
REGION Network 78: Sin requerimiento compresor 5
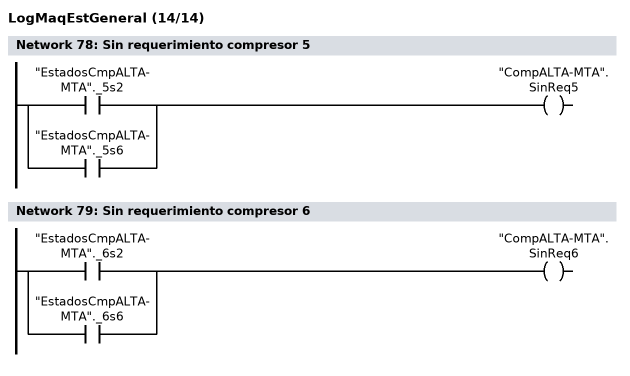
   RUNG wire#powerrail
      Contact( "EstadosCmpALTA-MTA"._5s2 )
      wire#w1
      Coil( "CompALTA-MTA".SinReq5 )
   END_RUNG
   RUNG wire#powerrail
      Contact( "EstadosCmpALTA-MTA"._5s6 )
   END_RUNG wire#w1
   // the same network as SCL:
   "CompALTA-MTA".SinReq5 := "EstadosCmpALTA-MTA"._5s2 OR "EstadosCmpALTA-MTA"._5s6;
END_REGION

REGION Network 79: Sin requerimiento compresor 6
   RUNG wire#powerrail
      Contact( "EstadosCmpALTA-MTA"._6s2 )
      wire#w1
      Coil( "CompALTA-MTA".SinReq6 )
   END_RUNG
   RUNG wire#powerrail
      Contact( "EstadosCmpALTA-MTA"._6s6 )
   END_RUNG wire#w1
   // the same network as SCL:
   "CompALTA-MTA".SinReq6 := "EstadosCmpALTA-MTA"._6s2 OR "EstadosCmpALTA-MTA"._6s6;
END_REGION
END_FUNCTION

FUNCTION "CalcEst1" : Void   // FC36, LAD
{ S7_Optimized_Access := 'FALSE' }
VERSION : 0.1
   VAR_TEMP   // added for the SCL form of the ladder/FBD networks
      _w1 : Bool;
   END_VAR
BEGIN

REGION Network 1
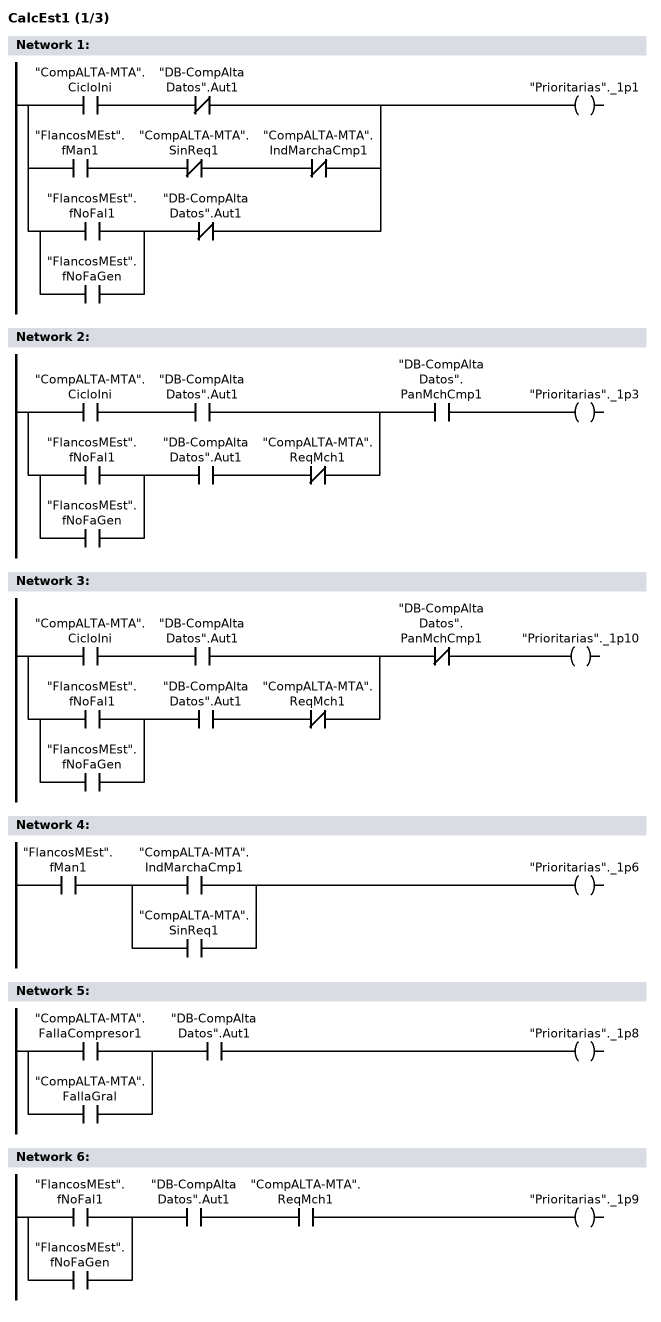
   RUNG wire#powerrail
      Contact( "CompALTA-MTA".CicloIni )
      I_Contact( "DB-CompAltaDatos".Aut1 )
      wire#w1
      Coil( "Prioritarias"._1p1 )
   END_RUNG
   RUNG wire#powerrail
      Contact( "FlancosMEst".fMan1 )
      I_Contact( "CompALTA-MTA".SinReq1 )
      I_Contact( "CompALTA-MTA".IndMarchaCmp1 )
   END_RUNG wire#w1
   RUNG wire#powerrail
      Contact( "FlancosMEst".fNoFal1 )
      wire#w2
      I_Contact( "DB-CompAltaDatos".Aut1 )
   END_RUNG wire#w1
   RUNG wire#powerrail
      Contact( "FlancosMEst".fNoFaGen )
   END_RUNG wire#w2
   // the same network as SCL:
   "Prioritarias"._1p1 := ("CompALTA-MTA".CicloIni AND NOT "DB-CompAltaDatos".Aut1) OR ("FlancosMEst".fMan1 AND NOT "CompALTA-MTA".SinReq1 AND NOT "CompALTA-MTA".IndMarchaCmp1) OR (("FlancosMEst".fNoFal1 OR "FlancosMEst".fNoFaGen) AND NOT "DB-CompAltaDatos".Aut1);
END_REGION

REGION Network 2
   RUNG wire#powerrail
      Contact( "CompALTA-MTA".CicloIni )
      Contact( "DB-CompAltaDatos".Aut1 )
      wire#w1
      Contact( "DB-CompAltaDatos".PanMchCmp1 )
      Coil( "Prioritarias"._1p3 )
   END_RUNG
   RUNG wire#powerrail
      Contact( "FlancosMEst".fNoFal1 )
      wire#w2
      Contact( "DB-CompAltaDatos".Aut1 )
      I_Contact( "CompALTA-MTA".ReqMch1 )
   END_RUNG wire#w1
   RUNG wire#powerrail
      Contact( "FlancosMEst".fNoFaGen )
   END_RUNG wire#w2
   // the same network as SCL:
   "Prioritarias"._1p3 := (("CompALTA-MTA".CicloIni AND "DB-CompAltaDatos".Aut1) OR (("FlancosMEst".fNoFal1 OR "FlancosMEst".fNoFaGen) AND "DB-CompAltaDatos".Aut1 AND NOT "CompALTA-MTA".ReqMch1)) AND "DB-CompAltaDatos".PanMchCmp1;
END_REGION

REGION Network 3
   RUNG wire#powerrail
      Contact( "CompALTA-MTA".CicloIni )
      Contact( "DB-CompAltaDatos".Aut1 )
      wire#w1
      I_Contact( "DB-CompAltaDatos".PanMchCmp1 )
      Coil( "Prioritarias"._1p10 )
   END_RUNG
   RUNG wire#powerrail
      Contact( "FlancosMEst".fNoFal1 )
      wire#w2
      Contact( "DB-CompAltaDatos".Aut1 )
      I_Contact( "CompALTA-MTA".ReqMch1 )
   END_RUNG wire#w1
   RUNG wire#powerrail
      Contact( "FlancosMEst".fNoFaGen )
   END_RUNG wire#w2
   // the same network as SCL:
   "Prioritarias"._1p10 := (("CompALTA-MTA".CicloIni AND "DB-CompAltaDatos".Aut1) OR (("FlancosMEst".fNoFal1 OR "FlancosMEst".fNoFaGen) AND "DB-CompAltaDatos".Aut1 AND NOT "CompALTA-MTA".ReqMch1)) AND NOT "DB-CompAltaDatos".PanMchCmp1;
END_REGION

REGION Network 4
   RUNG wire#powerrail
      Contact( "FlancosMEst".fMan1 )
      wire#w1
      Contact( "CompALTA-MTA".IndMarchaCmp1 )
      wire#w2
      Coil( "Prioritarias"._1p6 )
   END_RUNG
   RUNG wire#w1
      Contact( "CompALTA-MTA".SinReq1 )
   END_RUNG wire#w2
   // the same network as SCL:
   "Prioritarias"._1p6 := "FlancosMEst".fMan1 AND ("CompALTA-MTA".IndMarchaCmp1 OR "CompALTA-MTA".SinReq1);
END_REGION

REGION Network 5
   RUNG wire#powerrail
      Contact( "CompALTA-MTA".FallaCompresor1 )
      wire#w1
      Contact( "DB-CompAltaDatos".Aut1 )
      Coil( "Prioritarias"._1p8 )
   END_RUNG
   RUNG wire#powerrail
      Contact( "CompALTA-MTA".FallaGral )
   END_RUNG wire#w1
   // the same network as SCL:
   "Prioritarias"._1p8 := ("CompALTA-MTA".FallaCompresor1 OR "CompALTA-MTA".FallaGral) AND "DB-CompAltaDatos".Aut1;
END_REGION

REGION Network 6
   RUNG wire#powerrail
      Contact( "FlancosMEst".fNoFal1 )
      wire#w1
      Contact( "DB-CompAltaDatos".Aut1 )
      Contact( "CompALTA-MTA".ReqMch1 )
      Coil( "Prioritarias"._1p9 )
   END_RUNG
   RUNG wire#powerrail
      Contact( "FlancosMEst".fNoFaGen )
   END_RUNG wire#w1
   // the same network as SCL:
   "Prioritarias"._1p9 := ("FlancosMEst".fNoFal1 OR "FlancosMEst".fNoFaGen) AND "DB-CompAltaDatos".Aut1 AND "CompALTA-MTA".ReqMch1;
END_REGION

REGION Network 7
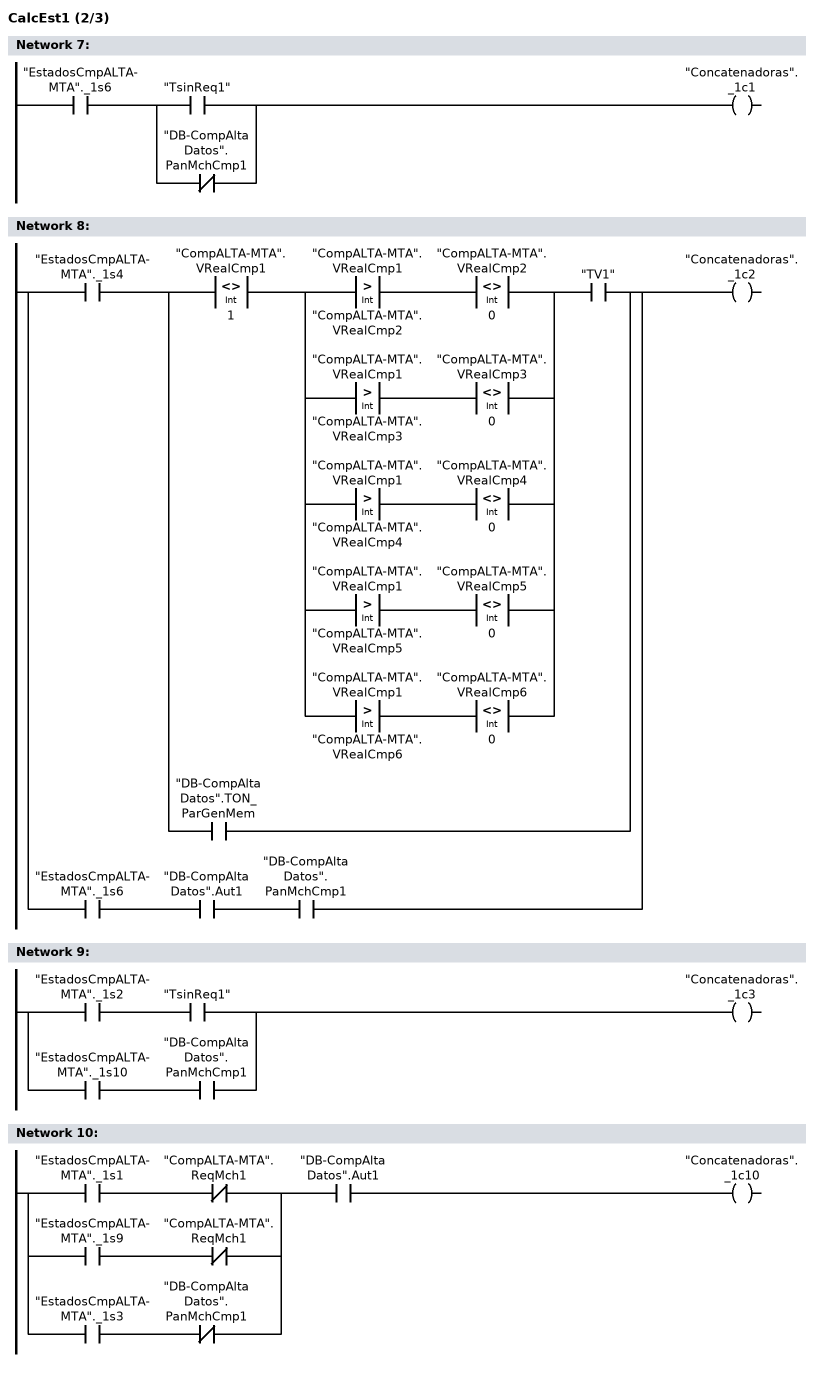
   RUNG wire#powerrail
      Contact( "EstadosCmpALTA-MTA"._1s6 )
      wire#w1
      Contact( "TsinReq1" )
      wire#w2
      Coil( "Concatenadoras"._1c1 )
   END_RUNG
   RUNG wire#w1
      I_Contact( "DB-CompAltaDatos".PanMchCmp1 )
   END_RUNG wire#w2
   // the same network as SCL:
   "Concatenadoras"._1c1 := "EstadosCmpALTA-MTA"._1s6 AND ("TsinReq1" OR NOT "DB-CompAltaDatos".PanMchCmp1);
END_REGION

REGION Network 8
   RUNG wire#powerrail
      Contact( "EstadosCmpALTA-MTA"._1s4 )
      wire#w1
      { S7_Templates := "SrcType := Int" } NE_Contact(in1 := "CompALTA-MTA".VRealCmp1, in2 := 1)
      wire#w2
      { S7_Templates := "SrcType := Int" } GT_Contact(in1 := "CompALTA-MTA".VRealCmp1, in2 := "CompALTA-MTA".VRealCmp2)
      { S7_Templates := "SrcType := Int" } NE_Contact(in1 := "CompALTA-MTA".VRealCmp2, in2 := 0)
      wire#w3
      Contact( "TV1" )
      wire#w4
      Coil( "Concatenadoras"._1c2 )
   END_RUNG
   RUNG wire#w2
      { S7_Templates := "SrcType := Int" } GT_Contact(in1 := "CompALTA-MTA".VRealCmp1, in2 := "CompALTA-MTA".VRealCmp3)
      { S7_Templates := "SrcType := Int" } NE_Contact(in1 := "CompALTA-MTA".VRealCmp3, in2 := 0)
   END_RUNG wire#w3
   RUNG wire#w2
      { S7_Templates := "SrcType := Int" } GT_Contact(in1 := "CompALTA-MTA".VRealCmp1, in2 := "CompALTA-MTA".VRealCmp4)
      { S7_Templates := "SrcType := Int" } NE_Contact(in1 := "CompALTA-MTA".VRealCmp4, in2 := 0)
   END_RUNG wire#w3
   RUNG wire#w2
      { S7_Templates := "SrcType := Int" } GT_Contact(in1 := "CompALTA-MTA".VRealCmp1, in2 := "CompALTA-MTA".VRealCmp5)
      { S7_Templates := "SrcType := Int" } NE_Contact(in1 := "CompALTA-MTA".VRealCmp5, in2 := 0)
   END_RUNG wire#w3
   RUNG wire#w2
      { S7_Templates := "SrcType := Int" } GT_Contact(in1 := "CompALTA-MTA".VRealCmp1, in2 := "CompALTA-MTA".VRealCmp6)
      { S7_Templates := "SrcType := Int" } NE_Contact(in1 := "CompALTA-MTA".VRealCmp6, in2 := 0)
   END_RUNG wire#w3
   RUNG wire#w1
      Contact( "DB-CompAltaDatos".TON_ParGenMem )
   END_RUNG wire#w4
   RUNG wire#powerrail
      Contact( "EstadosCmpALTA-MTA"._1s6 )
      Contact( "DB-CompAltaDatos".Aut1 )
      Contact( "DB-CompAltaDatos".PanMchCmp1 )
   END_RUNG wire#w4
   // the same network as SCL:
   "Concatenadoras"._1c2 := ("EstadosCmpALTA-MTA"._1s4 AND ((("CompALTA-MTA".VRealCmp1 <> 1) AND ((("CompALTA-MTA".VRealCmp1 > "CompALTA-MTA".VRealCmp2) AND ("CompALTA-MTA".VRealCmp2 <> 0)) OR (("CompALTA-MTA".VRealCmp1 > "CompALTA-MTA".VRealCmp3) AND ("CompALTA-MTA".VRealCmp3 <> 0)) OR (("CompALTA-MTA".VRealCmp1 > "CompALTA-MTA".VRealCmp4) AND ("CompALTA-MTA".VRealCmp4 <> 0)) OR (("CompALTA-MTA".VRealCmp1 > "CompALTA-MTA".VRealCmp5) AND ("CompALTA-MTA".VRealCmp5 <> 0)) OR (("CompALTA-MTA".VRealCmp1 > "CompALTA-MTA".VRealCmp6) AND ("CompALTA-MTA".VRealCmp6 <> 0))) AND "TV1") OR "DB-CompAltaDatos".TON_ParGenMem)) OR ("EstadosCmpALTA-MTA"._1s6 AND "DB-CompAltaDatos".Aut1 AND "DB-CompAltaDatos".PanMchCmp1);
END_REGION

REGION Network 9
   RUNG wire#powerrail
      Contact( "EstadosCmpALTA-MTA"._1s2 )
      Contact( "TsinReq1" )
      wire#w1
      Coil( "Concatenadoras"._1c3 )
   END_RUNG
   RUNG wire#powerrail
      Contact( "EstadosCmpALTA-MTA"._1s10 )
      Contact( "DB-CompAltaDatos".PanMchCmp1 )
   END_RUNG wire#w1
   // the same network as SCL:
   "Concatenadoras"._1c3 := ("EstadosCmpALTA-MTA"._1s2 AND "TsinReq1") OR ("EstadosCmpALTA-MTA"._1s10 AND "DB-CompAltaDatos".PanMchCmp1);
END_REGION

REGION Network 10
   RUNG wire#powerrail
      Contact( "EstadosCmpALTA-MTA"._1s1 )
      I_Contact( "CompALTA-MTA".ReqMch1 )
      wire#w1
      Contact( "DB-CompAltaDatos".Aut1 )
      Coil( "Concatenadoras"._1c10 )
   END_RUNG
   RUNG wire#powerrail
      Contact( "EstadosCmpALTA-MTA"._1s9 )
      I_Contact( "CompALTA-MTA".ReqMch1 )
   END_RUNG wire#w1
   RUNG wire#powerrail
      Contact( "EstadosCmpALTA-MTA"._1s3 )
      I_Contact( "DB-CompAltaDatos".PanMchCmp1 )
   END_RUNG wire#w1
   // the same network as SCL:
   "Concatenadoras"._1c10 := (("EstadosCmpALTA-MTA"._1s1 AND NOT "CompALTA-MTA".ReqMch1) OR ("EstadosCmpALTA-MTA"._1s9 AND NOT "CompALTA-MTA".ReqMch1) OR ("EstadosCmpALTA-MTA"._1s3 AND NOT "DB-CompAltaDatos".PanMchCmp1)) AND "DB-CompAltaDatos".Aut1;
END_REGION

REGION Network 11
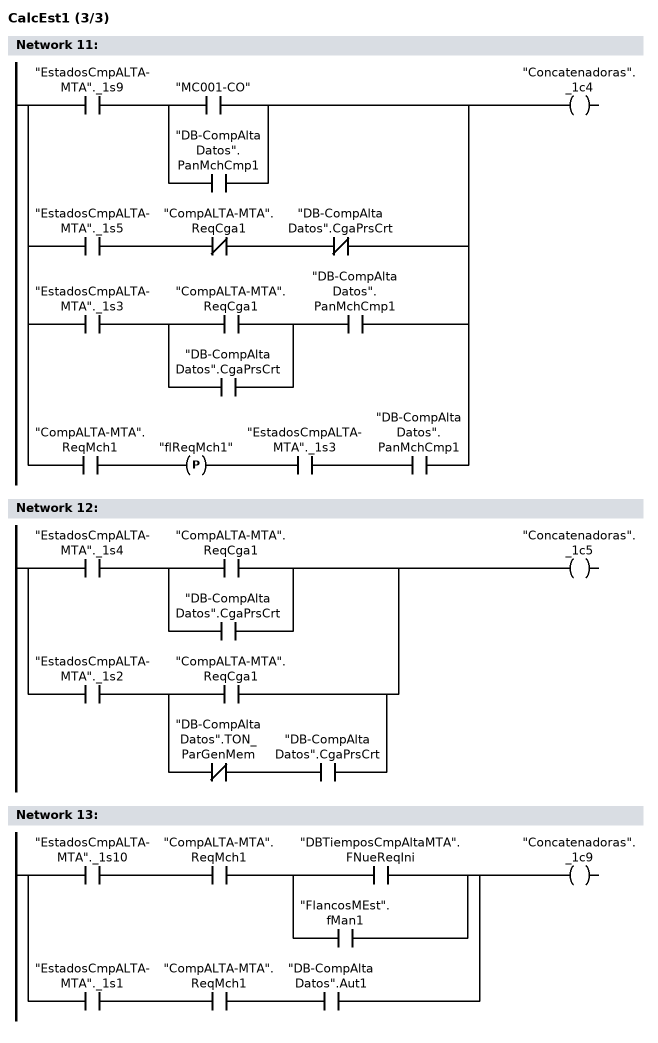
   RUNG wire#powerrail
      Contact( "EstadosCmpALTA-MTA"._1s9 )
      wire#w1
      Contact( "MC001-CO" )
      wire#w2
      Coil( "Concatenadoras"._1c4 )
   END_RUNG
   RUNG wire#w1
      Contact( "DB-CompAltaDatos".PanMchCmp1 )
   END_RUNG wire#w2
   RUNG wire#powerrail
      Contact( "EstadosCmpALTA-MTA"._1s5 )
      I_Contact( "CompALTA-MTA".ReqCga1 )
      I_Contact( "DB-CompAltaDatos".CgaPrsCrt )
   END_RUNG wire#w2
   RUNG wire#powerrail
      Contact( "EstadosCmpALTA-MTA"._1s3 )
      wire#w3
      Contact( "CompALTA-MTA".ReqCga1 )
      wire#w4
      Contact( "DB-CompAltaDatos".PanMchCmp1 )
   END_RUNG wire#w2
   RUNG wire#w3
      Contact( "DB-CompAltaDatos".CgaPrsCrt )
   END_RUNG wire#w4
   RUNG wire#powerrail
      Contact( "CompALTA-MTA".ReqMch1 )
      P_Trig( "flReqMch1" )
      Contact( "EstadosCmpALTA-MTA"._1s3 )
      Contact( "DB-CompAltaDatos".PanMchCmp1 )
   END_RUNG wire#w2
   // the same network as SCL:
   #_w1 := "CompALTA-MTA".ReqMch1 AND NOT "flReqMch1";   // rising edge
   "flReqMch1" := "CompALTA-MTA".ReqMch1;
   "Concatenadoras"._1c4 := ("EstadosCmpALTA-MTA"._1s9 AND ("MC001-CO" OR "DB-CompAltaDatos".PanMchCmp1)) OR ("EstadosCmpALTA-MTA"._1s5 AND NOT "CompALTA-MTA".ReqCga1 AND NOT "DB-CompAltaDatos".CgaPrsCrt) OR ("EstadosCmpALTA-MTA"._1s3 AND ("CompALTA-MTA".ReqCga1 OR "DB-CompAltaDatos".CgaPrsCrt) AND "DB-CompAltaDatos".PanMchCmp1) OR (#_w1 AND "EstadosCmpALTA-MTA"._1s3 AND "DB-CompAltaDatos".PanMchCmp1);
END_REGION

REGION Network 12
   RUNG wire#powerrail
      Contact( "EstadosCmpALTA-MTA"._1s4 )
      wire#w1
      Contact( "CompALTA-MTA".ReqCga1 )
      wire#w2
      Coil( "Concatenadoras"._1c5 )
   END_RUNG
   RUNG wire#w1
      Contact( "DB-CompAltaDatos".CgaPrsCrt )
   END_RUNG wire#w2
   RUNG wire#powerrail
      Contact( "EstadosCmpALTA-MTA"._1s2 )
      wire#w3
      Contact( "CompALTA-MTA".ReqCga1 )
   END_RUNG wire#w2
   RUNG wire#w3
      I_Contact( "DB-CompAltaDatos".TON_ParGenMem )
      Contact( "DB-CompAltaDatos".CgaPrsCrt )
   END_RUNG wire#w2
   // the same network as SCL:
   "Concatenadoras"._1c5 := ("EstadosCmpALTA-MTA"._1s4 AND ("CompALTA-MTA".ReqCga1 OR "DB-CompAltaDatos".CgaPrsCrt)) OR ("EstadosCmpALTA-MTA"._1s2 AND ("CompALTA-MTA".ReqCga1 OR (NOT "DB-CompAltaDatos".TON_ParGenMem AND "DB-CompAltaDatos".CgaPrsCrt)));
END_REGION

REGION Network 13
   RUNG wire#powerrail
      Contact( "EstadosCmpALTA-MTA"._1s10 )
      Contact( "CompALTA-MTA".ReqMch1 )
      wire#w1
      Contact( "DBTiemposCmpAltaMTA".FNueReqIni )
      wire#w2
      Coil( "Concatenadoras"._1c9 )
   END_RUNG
   RUNG wire#w1
      Contact( "FlancosMEst".fMan1 )
   END_RUNG wire#w2
   RUNG wire#powerrail
      Contact( "EstadosCmpALTA-MTA"._1s1 )
      Contact( "CompALTA-MTA".ReqMch1 )
      Contact( "DB-CompAltaDatos".Aut1 )
   END_RUNG wire#w2
   // the same network as SCL:
   "Concatenadoras"._1c9 := ("EstadosCmpALTA-MTA"._1s10 AND "CompALTA-MTA".ReqMch1 AND ("DBTiemposCmpAltaMTA".FNueReqIni OR "FlancosMEst".fMan1)) OR ("EstadosCmpALTA-MTA"._1s1 AND "CompALTA-MTA".ReqMch1 AND "DB-CompAltaDatos".Aut1);
END_REGION

REGION Network 14 (STL)
         CALL  "FC_MAQ_EST_16"
         ( IN0  := %DB127.DBW0,
           IN1  := %DB128.DBW0,
           OUT2 := "ErrPMQ1",
           OUT3 := "ErrCMQ1",
           IO4  := %DB120.DBW0
         );
         NOP   0;
END_REGION

REGION Network 15 (STL)
         CALL  "FC-ANIM-CMP"
         ( IN0  := %DB120.DBW0,
           OUT1 := "CompALTA-MTA".AnimCMP1
         );
         NOP   0;
END_REGION
END_FUNCTION

FUNCTION "CalcEst2" : Void   // FC37, LAD
{ S7_Optimized_Access := 'FALSE' }
VERSION : 0.1
   VAR_TEMP   // added for the SCL form of the ladder/FBD networks
      _w1 : Bool;
   END_VAR
BEGIN

REGION Network 1
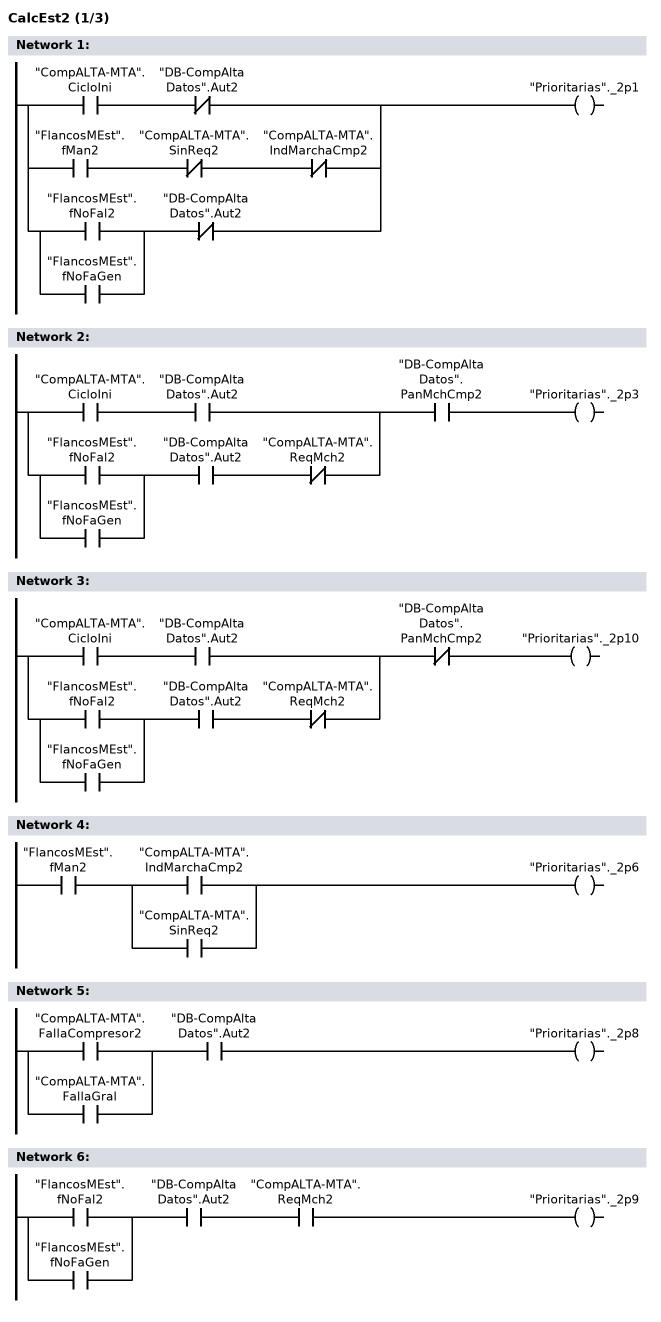
   RUNG wire#powerrail
      Contact( "CompALTA-MTA".CicloIni )
      I_Contact( "DB-CompAltaDatos".Aut2 )
      wire#w1
      Coil( "Prioritarias"._2p1 )
   END_RUNG
   RUNG wire#powerrail
      Contact( "FlancosMEst".fMan2 )
      I_Contact( "CompALTA-MTA".SinReq2 )
      I_Contact( "CompALTA-MTA".IndMarchaCmp2 )
   END_RUNG wire#w1
   RUNG wire#powerrail
      Contact( "FlancosMEst".fNoFal2 )
      wire#w2
      I_Contact( "DB-CompAltaDatos".Aut2 )
   END_RUNG wire#w1
   RUNG wire#powerrail
      Contact( "FlancosMEst".fNoFaGen )
   END_RUNG wire#w2
   // the same network as SCL:
   "Prioritarias"._2p1 := ("CompALTA-MTA".CicloIni AND NOT "DB-CompAltaDatos".Aut2) OR ("FlancosMEst".fMan2 AND NOT "CompALTA-MTA".SinReq2 AND NOT "CompALTA-MTA".IndMarchaCmp2) OR (("FlancosMEst".fNoFal2 OR "FlancosMEst".fNoFaGen) AND NOT "DB-CompAltaDatos".Aut2);
END_REGION

REGION Network 2
   RUNG wire#powerrail
      Contact( "CompALTA-MTA".CicloIni )
      Contact( "DB-CompAltaDatos".Aut2 )
      wire#w1
      Contact( "DB-CompAltaDatos".PanMchCmp2 )
      Coil( "Prioritarias"._2p3 )
   END_RUNG
   RUNG wire#powerrail
      Contact( "FlancosMEst".fNoFal2 )
      wire#w2
      Contact( "DB-CompAltaDatos".Aut2 )
      I_Contact( "CompALTA-MTA".ReqMch2 )
   END_RUNG wire#w1
   RUNG wire#powerrail
      Contact( "FlancosMEst".fNoFaGen )
   END_RUNG wire#w2
   // the same network as SCL:
   "Prioritarias"._2p3 := (("CompALTA-MTA".CicloIni AND "DB-CompAltaDatos".Aut2) OR (("FlancosMEst".fNoFal2 OR "FlancosMEst".fNoFaGen) AND "DB-CompAltaDatos".Aut2 AND NOT "CompALTA-MTA".ReqMch2)) AND "DB-CompAltaDatos".PanMchCmp2;
END_REGION

REGION Network 3
   RUNG wire#powerrail
      Contact( "CompALTA-MTA".CicloIni )
      Contact( "DB-CompAltaDatos".Aut2 )
      wire#w1
      I_Contact( "DB-CompAltaDatos".PanMchCmp2 )
      Coil( "Prioritarias"._2p10 )
   END_RUNG
   RUNG wire#powerrail
      Contact( "FlancosMEst".fNoFal2 )
      wire#w2
      Contact( "DB-CompAltaDatos".Aut2 )
      I_Contact( "CompALTA-MTA".ReqMch2 )
   END_RUNG wire#w1
   RUNG wire#powerrail
      Contact( "FlancosMEst".fNoFaGen )
   END_RUNG wire#w2
   // the same network as SCL:
   "Prioritarias"._2p10 := (("CompALTA-MTA".CicloIni AND "DB-CompAltaDatos".Aut2) OR (("FlancosMEst".fNoFal2 OR "FlancosMEst".fNoFaGen) AND "DB-CompAltaDatos".Aut2 AND NOT "CompALTA-MTA".ReqMch2)) AND NOT "DB-CompAltaDatos".PanMchCmp2;
END_REGION

REGION Network 4
   RUNG wire#powerrail
      Contact( "FlancosMEst".fMan2 )
      wire#w1
      Contact( "CompALTA-MTA".IndMarchaCmp2 )
      wire#w2
      Coil( "Prioritarias"._2p6 )
   END_RUNG
   RUNG wire#w1
      Contact( "CompALTA-MTA".SinReq2 )
   END_RUNG wire#w2
   // the same network as SCL:
   "Prioritarias"._2p6 := "FlancosMEst".fMan2 AND ("CompALTA-MTA".IndMarchaCmp2 OR "CompALTA-MTA".SinReq2);
END_REGION

REGION Network 5
   RUNG wire#powerrail
      Contact( "CompALTA-MTA".FallaCompresor2 )
      wire#w1
      Contact( "DB-CompAltaDatos".Aut2 )
      Coil( "Prioritarias"._2p8 )
   END_RUNG
   RUNG wire#powerrail
      Contact( "CompALTA-MTA".FallaGral )
   END_RUNG wire#w1
   // the same network as SCL:
   "Prioritarias"._2p8 := ("CompALTA-MTA".FallaCompresor2 OR "CompALTA-MTA".FallaGral) AND "DB-CompAltaDatos".Aut2;
END_REGION

REGION Network 6
   RUNG wire#powerrail
      Contact( "FlancosMEst".fNoFal2 )
      wire#w1
      Contact( "DB-CompAltaDatos".Aut2 )
      Contact( "CompALTA-MTA".ReqMch2 )
      Coil( "Prioritarias"._2p9 )
   END_RUNG
   RUNG wire#powerrail
      Contact( "FlancosMEst".fNoFaGen )
   END_RUNG wire#w1
   // the same network as SCL:
   "Prioritarias"._2p9 := ("FlancosMEst".fNoFal2 OR "FlancosMEst".fNoFaGen) AND "DB-CompAltaDatos".Aut2 AND "CompALTA-MTA".ReqMch2;
END_REGION

REGION Network 7
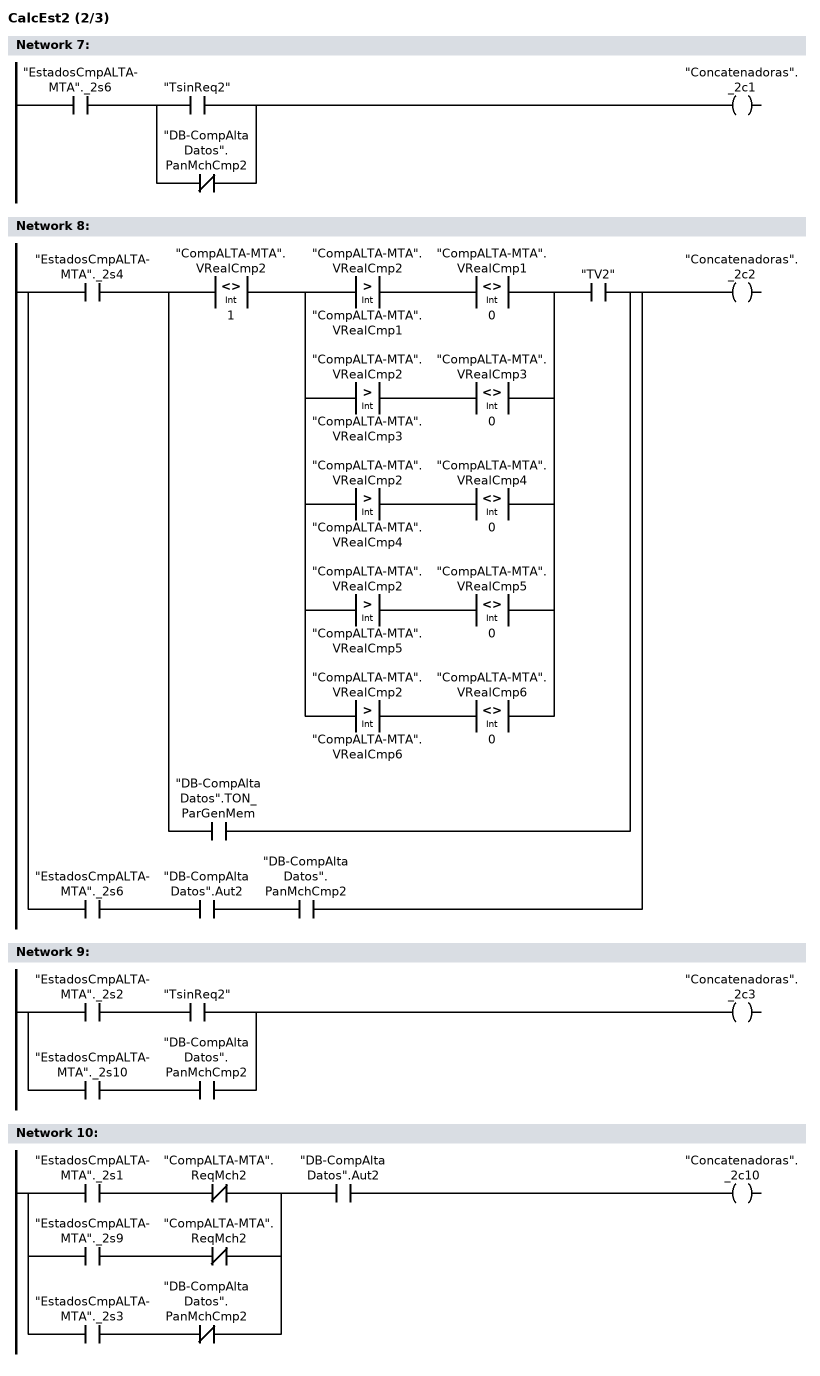
   RUNG wire#powerrail
      Contact( "EstadosCmpALTA-MTA"._2s6 )
      wire#w1
      Contact( "TsinReq2" )
      wire#w2
      Coil( "Concatenadoras"._2c1 )
   END_RUNG
   RUNG wire#w1
      I_Contact( "DB-CompAltaDatos".PanMchCmp2 )
   END_RUNG wire#w2
   // the same network as SCL:
   "Concatenadoras"._2c1 := "EstadosCmpALTA-MTA"._2s6 AND ("TsinReq2" OR NOT "DB-CompAltaDatos".PanMchCmp2);
END_REGION

REGION Network 8
   RUNG wire#powerrail
      Contact( "EstadosCmpALTA-MTA"._2s4 )
      wire#w1
      { S7_Templates := "SrcType := Int" } NE_Contact(in1 := "CompALTA-MTA".VRealCmp2, in2 := 1)
      wire#w2
      { S7_Templates := "SrcType := Int" } GT_Contact(in1 := "CompALTA-MTA".VRealCmp2, in2 := "CompALTA-MTA".VRealCmp1)
      { S7_Templates := "SrcType := Int" } NE_Contact(in1 := "CompALTA-MTA".VRealCmp1, in2 := 0)
      wire#w3
      Contact( "TV2" )
      wire#w4
      Coil( "Concatenadoras"._2c2 )
   END_RUNG
   RUNG wire#w2
      { S7_Templates := "SrcType := Int" } GT_Contact(in1 := "CompALTA-MTA".VRealCmp2, in2 := "CompALTA-MTA".VRealCmp3)
      { S7_Templates := "SrcType := Int" } NE_Contact(in1 := "CompALTA-MTA".VRealCmp3, in2 := 0)
   END_RUNG wire#w3
   RUNG wire#w2
      { S7_Templates := "SrcType := Int" } GT_Contact(in1 := "CompALTA-MTA".VRealCmp2, in2 := "CompALTA-MTA".VRealCmp4)
      { S7_Templates := "SrcType := Int" } NE_Contact(in1 := "CompALTA-MTA".VRealCmp4, in2 := 0)
   END_RUNG wire#w3
   RUNG wire#w2
      { S7_Templates := "SrcType := Int" } GT_Contact(in1 := "CompALTA-MTA".VRealCmp2, in2 := "CompALTA-MTA".VRealCmp5)
      { S7_Templates := "SrcType := Int" } NE_Contact(in1 := "CompALTA-MTA".VRealCmp5, in2 := 0)
   END_RUNG wire#w3
   RUNG wire#w2
      { S7_Templates := "SrcType := Int" } GT_Contact(in1 := "CompALTA-MTA".VRealCmp2, in2 := "CompALTA-MTA".VRealCmp6)
      { S7_Templates := "SrcType := Int" } NE_Contact(in1 := "CompALTA-MTA".VRealCmp6, in2 := 0)
   END_RUNG wire#w3
   RUNG wire#w1
      Contact( "DB-CompAltaDatos".TON_ParGenMem )
   END_RUNG wire#w4
   RUNG wire#powerrail
      Contact( "EstadosCmpALTA-MTA"._2s6 )
      Contact( "DB-CompAltaDatos".Aut2 )
      Contact( "DB-CompAltaDatos".PanMchCmp2 )
   END_RUNG wire#w4
   // the same network as SCL:
   "Concatenadoras"._2c2 := ("EstadosCmpALTA-MTA"._2s4 AND ((("CompALTA-MTA".VRealCmp2 <> 1) AND ((("CompALTA-MTA".VRealCmp2 > "CompALTA-MTA".VRealCmp1) AND ("CompALTA-MTA".VRealCmp1 <> 0)) OR (("CompALTA-MTA".VRealCmp2 > "CompALTA-MTA".VRealCmp3) AND ("CompALTA-MTA".VRealCmp3 <> 0)) OR (("CompALTA-MTA".VRealCmp2 > "CompALTA-MTA".VRealCmp4) AND ("CompALTA-MTA".VRealCmp4 <> 0)) OR (("CompALTA-MTA".VRealCmp2 > "CompALTA-MTA".VRealCmp5) AND ("CompALTA-MTA".VRealCmp5 <> 0)) OR (("CompALTA-MTA".VRealCmp2 > "CompALTA-MTA".VRealCmp6) AND ("CompALTA-MTA".VRealCmp6 <> 0))) AND "TV2") OR "DB-CompAltaDatos".TON_ParGenMem)) OR ("EstadosCmpALTA-MTA"._2s6 AND "DB-CompAltaDatos".Aut2 AND "DB-CompAltaDatos".PanMchCmp2);
END_REGION

REGION Network 9
   RUNG wire#powerrail
      Contact( "EstadosCmpALTA-MTA"._2s2 )
      Contact( "TsinReq2" )
      wire#w1
      Coil( "Concatenadoras"._2c3 )
   END_RUNG
   RUNG wire#powerrail
      Contact( "EstadosCmpALTA-MTA"._2s10 )
      Contact( "DB-CompAltaDatos".PanMchCmp2 )
   END_RUNG wire#w1
   // the same network as SCL:
   "Concatenadoras"._2c3 := ("EstadosCmpALTA-MTA"._2s2 AND "TsinReq2") OR ("EstadosCmpALTA-MTA"._2s10 AND "DB-CompAltaDatos".PanMchCmp2);
END_REGION

REGION Network 10
   RUNG wire#powerrail
      Contact( "EstadosCmpALTA-MTA"._2s1 )
      I_Contact( "CompALTA-MTA".ReqMch2 )
      wire#w1
      Contact( "DB-CompAltaDatos".Aut2 )
      Coil( "Concatenadoras"._2c10 )
   END_RUNG
   RUNG wire#powerrail
      Contact( "EstadosCmpALTA-MTA"._2s9 )
      I_Contact( "CompALTA-MTA".ReqMch2 )
   END_RUNG wire#w1
   RUNG wire#powerrail
      Contact( "EstadosCmpALTA-MTA"._2s3 )
      I_Contact( "DB-CompAltaDatos".PanMchCmp2 )
   END_RUNG wire#w1
   // the same network as SCL:
   "Concatenadoras"._2c10 := (("EstadosCmpALTA-MTA"._2s1 AND NOT "CompALTA-MTA".ReqMch2) OR ("EstadosCmpALTA-MTA"._2s9 AND NOT "CompALTA-MTA".ReqMch2) OR ("EstadosCmpALTA-MTA"._2s3 AND NOT "DB-CompAltaDatos".PanMchCmp2)) AND "DB-CompAltaDatos".Aut2;
END_REGION

REGION Network 11
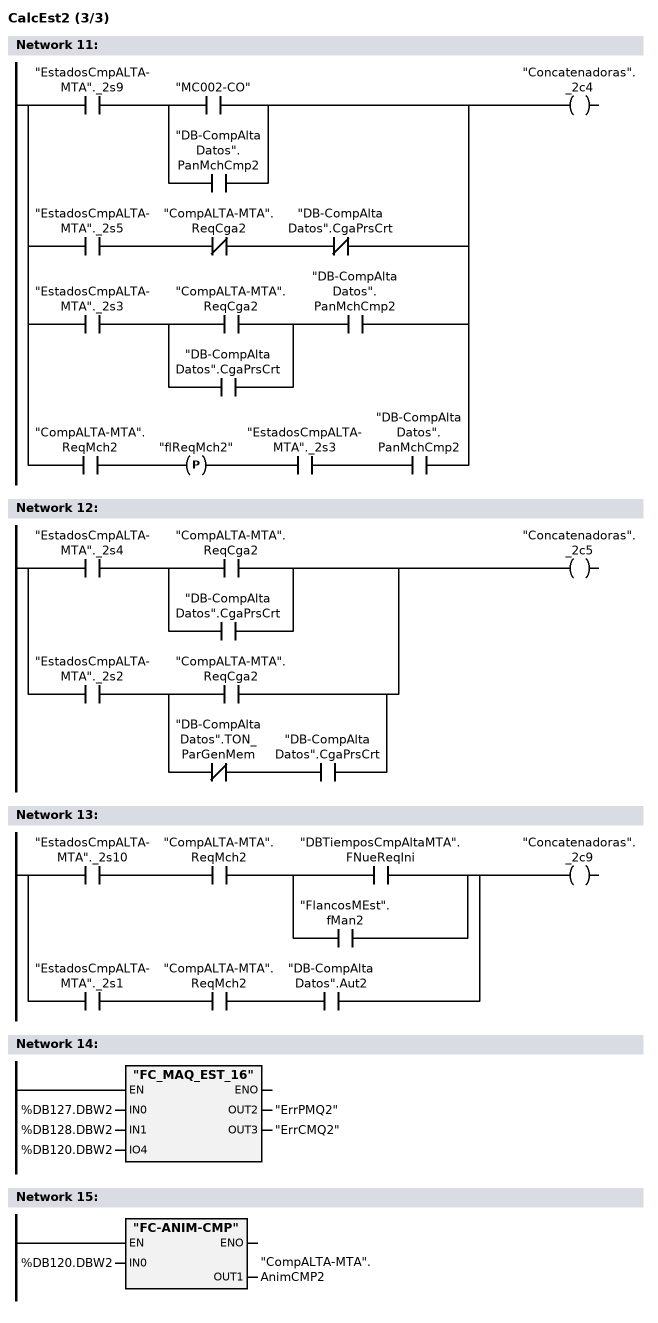
   RUNG wire#powerrail
      Contact( "EstadosCmpALTA-MTA"._2s9 )
      wire#w1
      Contact( "MC002-CO" )
      wire#w2
      Coil( "Concatenadoras"._2c4 )
   END_RUNG
   RUNG wire#w1
      Contact( "DB-CompAltaDatos".PanMchCmp2 )
   END_RUNG wire#w2
   RUNG wire#powerrail
      Contact( "EstadosCmpALTA-MTA"._2s5 )
      I_Contact( "CompALTA-MTA".ReqCga2 )
      I_Contact( "DB-CompAltaDatos".CgaPrsCrt )
   END_RUNG wire#w2
   RUNG wire#powerrail
      Contact( "EstadosCmpALTA-MTA"._2s3 )
      wire#w3
      Contact( "CompALTA-MTA".ReqCga2 )
      wire#w4
      Contact( "DB-CompAltaDatos".PanMchCmp2 )
   END_RUNG wire#w2
   RUNG wire#w3
      Contact( "DB-CompAltaDatos".CgaPrsCrt )
   END_RUNG wire#w4
   RUNG wire#powerrail
      Contact( "CompALTA-MTA".ReqMch2 )
      P_Trig( "flReqMch2" )
      Contact( "EstadosCmpALTA-MTA"._2s3 )
      Contact( "DB-CompAltaDatos".PanMchCmp2 )
   END_RUNG wire#w2
   // the same network as SCL:
   #_w1 := "CompALTA-MTA".ReqMch2 AND NOT "flReqMch2";   // rising edge
   "flReqMch2" := "CompALTA-MTA".ReqMch2;
   "Concatenadoras"._2c4 := ("EstadosCmpALTA-MTA"._2s9 AND ("MC002-CO" OR "DB-CompAltaDatos".PanMchCmp2)) OR ("EstadosCmpALTA-MTA"._2s5 AND NOT "CompALTA-MTA".ReqCga2 AND NOT "DB-CompAltaDatos".CgaPrsCrt) OR ("EstadosCmpALTA-MTA"._2s3 AND ("CompALTA-MTA".ReqCga2 OR "DB-CompAltaDatos".CgaPrsCrt) AND "DB-CompAltaDatos".PanMchCmp2) OR (#_w1 AND "EstadosCmpALTA-MTA"._2s3 AND "DB-CompAltaDatos".PanMchCmp2);
END_REGION

REGION Network 12
   RUNG wire#powerrail
      Contact( "EstadosCmpALTA-MTA"._2s4 )
      wire#w1
      Contact( "CompALTA-MTA".ReqCga2 )
      wire#w2
      Coil( "Concatenadoras"._2c5 )
   END_RUNG
   RUNG wire#w1
      Contact( "DB-CompAltaDatos".CgaPrsCrt )
   END_RUNG wire#w2
   RUNG wire#powerrail
      Contact( "EstadosCmpALTA-MTA"._2s2 )
      wire#w3
      Contact( "CompALTA-MTA".ReqCga2 )
   END_RUNG wire#w2
   RUNG wire#w3
      I_Contact( "DB-CompAltaDatos".TON_ParGenMem )
      Contact( "DB-CompAltaDatos".CgaPrsCrt )
   END_RUNG wire#w2
   // the same network as SCL:
   "Concatenadoras"._2c5 := ("EstadosCmpALTA-MTA"._2s4 AND ("CompALTA-MTA".ReqCga2 OR "DB-CompAltaDatos".CgaPrsCrt)) OR ("EstadosCmpALTA-MTA"._2s2 AND ("CompALTA-MTA".ReqCga2 OR (NOT "DB-CompAltaDatos".TON_ParGenMem AND "DB-CompAltaDatos".CgaPrsCrt)));
END_REGION

REGION Network 13
   RUNG wire#powerrail
      Contact( "EstadosCmpALTA-MTA"._2s10 )
      Contact( "CompALTA-MTA".ReqMch2 )
      wire#w1
      Contact( "DBTiemposCmpAltaMTA".FNueReqIni )
      wire#w2
      Coil( "Concatenadoras"._2c9 )
   END_RUNG
   RUNG wire#w1
      Contact( "FlancosMEst".fMan2 )
   END_RUNG wire#w2
   RUNG wire#powerrail
      Contact( "EstadosCmpALTA-MTA"._2s1 )
      Contact( "CompALTA-MTA".ReqMch2 )
      Contact( "DB-CompAltaDatos".Aut2 )
   END_RUNG wire#w2
   // the same network as SCL:
   "Concatenadoras"._2c9 := ("EstadosCmpALTA-MTA"._2s10 AND "CompALTA-MTA".ReqMch2 AND ("DBTiemposCmpAltaMTA".FNueReqIni OR "FlancosMEst".fMan2)) OR ("EstadosCmpALTA-MTA"._2s1 AND "CompALTA-MTA".ReqMch2 AND "DB-CompAltaDatos".Aut2);
END_REGION

REGION Network 14
   RUNG wire#powerrail
      "FC_MAQ_EST_16"(IN0 := %DB127.DBW2, IN1 := %DB128.DBW2, OUT2 => "ErrPMQ2", OUT3 => "ErrCMQ2", IO4 := %DB120.DBW2)
   END_RUNG
   // the same network as SCL:
   "FC_MAQ_EST_16"(IN0 := %DB127.DBW2,
                   IN1 := %DB128.DBW2,
                   IO4 := %DB120.DBW2,
                   OUT2 => "ErrPMQ2",
                   OUT3 => "ErrCMQ2");
END_REGION

REGION Network 15
   RUNG wire#powerrail
      "FC-ANIM-CMP"(IN0 := %DB120.DBW2, OUT1 => "CompALTA-MTA".AnimCMP2)
   END_RUNG
   // the same network as SCL:
   "FC-ANIM-CMP"(IN0 := %DB120.DBW2, OUT1 => "CompALTA-MTA".AnimCMP2);
END_REGION
END_FUNCTION

FUNCTION "CalcEst3" : Void   // FC38, LAD
{ S7_Optimized_Access := 'FALSE' }
VERSION : 0.1
   VAR_TEMP   // added for the SCL form of the ladder/FBD networks
      _w1 : Bool;
   END_VAR
BEGIN

REGION Network 1
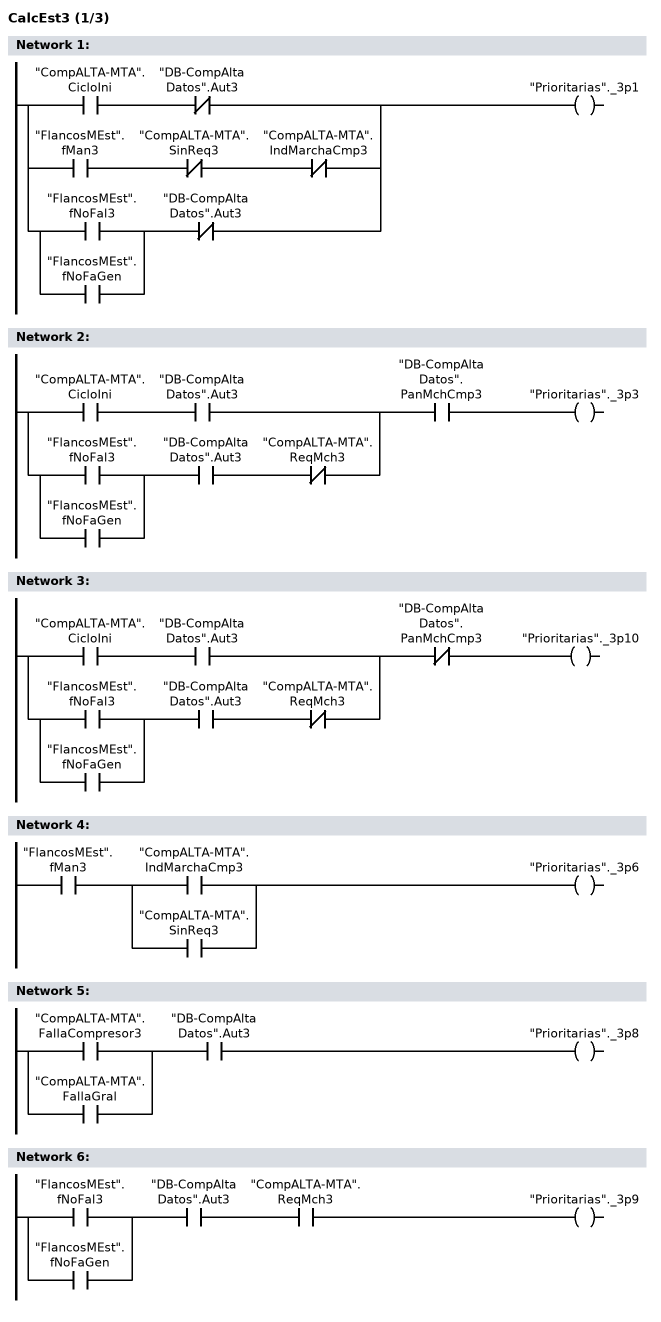
   RUNG wire#powerrail
      Contact( "CompALTA-MTA".CicloIni )
      I_Contact( "DB-CompAltaDatos".Aut3 )
      wire#w1
      Coil( "Prioritarias"._3p1 )
   END_RUNG
   RUNG wire#powerrail
      Contact( "FlancosMEst".fMan3 )
      I_Contact( "CompALTA-MTA".SinReq3 )
      I_Contact( "CompALTA-MTA".IndMarchaCmp3 )
   END_RUNG wire#w1
   RUNG wire#powerrail
      Contact( "FlancosMEst".fNoFal3 )
      wire#w2
      I_Contact( "DB-CompAltaDatos".Aut3 )
   END_RUNG wire#w1
   RUNG wire#powerrail
      Contact( "FlancosMEst".fNoFaGen )
   END_RUNG wire#w2
   // the same network as SCL:
   "Prioritarias"._3p1 := ("CompALTA-MTA".CicloIni AND NOT "DB-CompAltaDatos".Aut3) OR ("FlancosMEst".fMan3 AND NOT "CompALTA-MTA".SinReq3 AND NOT "CompALTA-MTA".IndMarchaCmp3) OR (("FlancosMEst".fNoFal3 OR "FlancosMEst".fNoFaGen) AND NOT "DB-CompAltaDatos".Aut3);
END_REGION

REGION Network 2
   RUNG wire#powerrail
      Contact( "CompALTA-MTA".CicloIni )
      Contact( "DB-CompAltaDatos".Aut3 )
      wire#w1
      Contact( "DB-CompAltaDatos".PanMchCmp3 )
      Coil( "Prioritarias"._3p3 )
   END_RUNG
   RUNG wire#powerrail
      Contact( "FlancosMEst".fNoFal3 )
      wire#w2
      Contact( "DB-CompAltaDatos".Aut3 )
      I_Contact( "CompALTA-MTA".ReqMch3 )
   END_RUNG wire#w1
   RUNG wire#powerrail
      Contact( "FlancosMEst".fNoFaGen )
   END_RUNG wire#w2
   // the same network as SCL:
   "Prioritarias"._3p3 := (("CompALTA-MTA".CicloIni AND "DB-CompAltaDatos".Aut3) OR (("FlancosMEst".fNoFal3 OR "FlancosMEst".fNoFaGen) AND "DB-CompAltaDatos".Aut3 AND NOT "CompALTA-MTA".ReqMch3)) AND "DB-CompAltaDatos".PanMchCmp3;
END_REGION

REGION Network 3
   RUNG wire#powerrail
      Contact( "CompALTA-MTA".CicloIni )
      Contact( "DB-CompAltaDatos".Aut3 )
      wire#w1
      I_Contact( "DB-CompAltaDatos".PanMchCmp3 )
      Coil( "Prioritarias"._3p10 )
   END_RUNG
   RUNG wire#powerrail
      Contact( "FlancosMEst".fNoFal3 )
      wire#w2
      Contact( "DB-CompAltaDatos".Aut3 )
      I_Contact( "CompALTA-MTA".ReqMch3 )
   END_RUNG wire#w1
   RUNG wire#powerrail
      Contact( "FlancosMEst".fNoFaGen )
   END_RUNG wire#w2
   // the same network as SCL:
   "Prioritarias"._3p10 := (("CompALTA-MTA".CicloIni AND "DB-CompAltaDatos".Aut3) OR (("FlancosMEst".fNoFal3 OR "FlancosMEst".fNoFaGen) AND "DB-CompAltaDatos".Aut3 AND NOT "CompALTA-MTA".ReqMch3)) AND NOT "DB-CompAltaDatos".PanMchCmp3;
END_REGION

REGION Network 4
   RUNG wire#powerrail
      Contact( "FlancosMEst".fMan3 )
      wire#w1
      Contact( "CompALTA-MTA".IndMarchaCmp3 )
      wire#w2
      Coil( "Prioritarias"._3p6 )
   END_RUNG
   RUNG wire#w1
      Contact( "CompALTA-MTA".SinReq3 )
   END_RUNG wire#w2
   // the same network as SCL:
   "Prioritarias"._3p6 := "FlancosMEst".fMan3 AND ("CompALTA-MTA".IndMarchaCmp3 OR "CompALTA-MTA".SinReq3);
END_REGION

REGION Network 5
   RUNG wire#powerrail
      Contact( "CompALTA-MTA".FallaCompresor3 )
      wire#w1
      Contact( "DB-CompAltaDatos".Aut3 )
      Coil( "Prioritarias"._3p8 )
   END_RUNG
   RUNG wire#powerrail
      Contact( "CompALTA-MTA".FallaGral )
   END_RUNG wire#w1
   // the same network as SCL:
   "Prioritarias"._3p8 := ("CompALTA-MTA".FallaCompresor3 OR "CompALTA-MTA".FallaGral) AND "DB-CompAltaDatos".Aut3;
END_REGION

REGION Network 6
   RUNG wire#powerrail
      Contact( "FlancosMEst".fNoFal3 )
      wire#w1
      Contact( "DB-CompAltaDatos".Aut3 )
      Contact( "CompALTA-MTA".ReqMch3 )
      Coil( "Prioritarias"._3p9 )
   END_RUNG
   RUNG wire#powerrail
      Contact( "FlancosMEst".fNoFaGen )
   END_RUNG wire#w1
   // the same network as SCL:
   "Prioritarias"._3p9 := ("FlancosMEst".fNoFal3 OR "FlancosMEst".fNoFaGen) AND "DB-CompAltaDatos".Aut3 AND "CompALTA-MTA".ReqMch3;
END_REGION

REGION Network 7